VAR_GLOBAL   // PLC tag table "默认变量表"
   "送煤皮带备妥" AT %I0.0 : Bool;
   "送煤皮带运行" AT %I0.1 : Bool;
   "送煤皮带故障" AT %I0.2 : Bool;
   "除铁器备妥" AT %I0.3 : Bool;
   "除铁器运行" AT %I0.4 : Bool;
   "除铁器故障" AT %I0.5 : Bool;
   "定量给煤机备妥" AT %I0.6 : Bool;
   "定量给煤机运行" AT %I0.7 : Bool;
   "定量给煤机故障" AT %I1.0 : Bool;
   "煤粉收尘器备妥" AT %I1.1 : Bool;
   "煤粉收尘器运行" AT %I1.2 : Bool;
   "煤粉收尘器故障" AT %I1.3 : Bool;
   "立磨尾排风机远程" AT %I1.4 : Bool;
   "立磨尾排风机运行" AT %I1.5 : Bool;
   "立磨尾排风机故障" AT %I1.6 : Bool;
   "立磨尾排风机待机" AT %I1.7 : Bool;
   "立磨尾排高压柜远程" AT %I2.0 : Bool;
   "立磨尾排高压柜合闸" AT %I2.1 : Bool;
   "立磨尾排高压柜分闸" AT %I2.2 : Bool;
   "定量给煤机断料信号" AT %I2.3 : Bool;
   "定量给煤机左跑偏信号" AT %I2.4 : Bool;
   "定量给煤机右跑偏信号" AT %I2.5 : Bool;
   "给煤机断链信号" AT %I2.6 : Bool;
   "立磨给煤机累计脉冲" AT %I2.7 : Bool;
   "定量给料机远程" AT %I3.0 : Bool;
   "1#铰刀运行" AT %I3.1 : Bool;
   "2#铰刀运行" AT %I3.2 : Bool;
   "1#分割轮运行" AT %I3.3 : Bool;
   "2#分割轮运行" AT %I3.4 : Bool;
   "3#分割轮运行" AT %I3.5 : Bool;
   "4#分割轮运行" AT %I3.6 : Bool;
   "5#分割轮运行" AT %I3.7 : Bool;
   "立磨主机高压柜远程" AT %I4.0 : Bool;
   "立磨主机高压柜合闸" AT %I4.1 : Bool;
   "立磨主机高压柜分闸" AT %I4.2 : Bool;
   "立磨主机运行" AT %I4.3 : Bool;
   "立磨主机故障" AT %I4.4 : Bool;
   "允许主机启动" AT %I4.5 : Bool;
   "跳停主机" AT %I4.6 : Bool;
   "6#分割轮运行" AT %I5.0 : Bool;
   "7#分割轮运行" AT %I5.1 : Bool;
   "8#分割轮运行" AT %I5.2 : Bool;
   "9#分割轮运行" AT %I5.3 : Bool;
   "10#分割轮运行" AT %I5.4 : Bool;
   "立磨尾排风机水平震动1" AT %IW256 : Int;
   "立磨尾排风机水平震动2" AT %IW258 : Int;
   "立磨尾排风机垂直震动1" AT %IW260 : Int;
   "立磨尾排风机垂直震动2" AT %IW262 : Int;
   "立磨尾排风机入口压力1" AT %IW264 : Int;
   "立磨尾排风机入口压力2" AT %IW266 : Int;
   "立磨尾排风机出口压力1" AT %IW268 : Int;
   "尾排风机入口执行器反馈" AT %IW270 : Int;
   "立磨1#煤粉仓负压" AT %IW272 : Int;
   "立磨2#煤粉仓负压" AT %IW274 : Int;
   "立磨热风管道负压" AT %IW276 : Int;
   "立磨主电机运行电流" AT %IW278 : Int;
   "立磨给煤机流量" AT %IW280 : Int;
   "立磨出口压力1" AT %IW282 : Int;
   "立磨出口压力2" AT %IW284 : Int;
   "立磨尾排风机运行转速" AT %IW288 : Int;
   "立磨尾排风机运行电流" AT %IW290 : Int;
   "立磨尾排风机出口温度1" AT %IW292 : Int;
   "立磨尾排风机入口温度1" AT %IW296 : Int;
   "立磨尾排风机入口温度2" AT %IW298 : Int;
   "立磨入磨口温度" AT %IW300 : Int;
   "1#煤粉仓1#温度" AT %ID304 : DWord;
   "1#煤粉仓2#温度" AT %ID308 : DWord;
   "1#煤粉仓3#温度" AT %ID312 : DWord;
   "1#煤粉仓4#温度" AT %ID316 : DWord;
   "1#煤粉仓5#温度" AT %ID320 : DWord;
   "1#煤粉仓6#温度" AT %ID324 : DWord;
   "2#煤粉仓1#温度" AT %ID328 : DWord;
   "2#煤粉仓2#温度" AT %ID332 : DWord;
   "2#煤粉仓3#温度" AT %ID336 : DWord;
   "2#煤粉仓4#温度" AT %ID340 : DWord;
   "2#煤粉仓5#温度" AT %ID344 : DWord;
   "2#煤粉仓6#温度" AT %ID348 : DWord;
   "立磨机出口温度1" AT %ID352 : DWord;
   "立磨机出口温度2" AT %ID356 : DWord;
   "PID360" AT %ID360 : DWord;
   "PID364" AT %ID364 : DWord;
   "电机绕组U相温度" AT %ID368 : DWord;
   "电机绕组V相温度" AT %ID372 : DWord;
   "电机绕组W相温度" AT %ID376 : DWord;
   "尾排电机前轴温度" AT %ID380 : DWord;
   "尾排电机后轴温度" AT %ID384 : DWord;
   "尾排风机前轴温度" AT %ID388 : DWord;
   "尾排风机后轴温度" AT %ID392 : DWord;
   "PID396" AT %ID396 : DWord;
   "立磨主机远程" AT %I4.7 : Bool;
   "11#分割轮运行" AT %I5.5 : Bool;
   "12#分割轮运行" AT %I5.6 : Bool;
   "立磨主电机轻故障" AT %I5.7 : Bool;
   "1#板式给煤机-褐煤备妥" AT %I6.0 : Bool;
   "1#板式给煤机-褐煤运行" AT %I6.1 : Bool;
   "1#板式给煤机-褐煤故障" AT %I6.2 : Bool;
   "2#板式给煤机-烟煤备妥" AT %I6.3 : Bool;
   "2#板式给煤机-烟煤运行" AT %I6.4 : Bool;
   "2#板式给煤机-烟煤故障" AT %I6.5 : Bool;
   "1#板式给煤机-褐煤脉冲累计" AT %I6.6 : Bool;
   "2#板式给煤机-烟煤脉冲累计" AT %I6.7 : Bool;
   "储气罐阀门远程" AT %I7.0 : Bool;
   "储气罐阀门开到位" AT %I7.1 : Bool;
   "储气罐阀门关到位" AT %I7.2 : Bool;
   "I7_3" AT %I7.3 : Bool;
   "I7_4" AT %I7.4 : Bool;
   "I7_5" AT %I7.5 : Bool;
   "I7_6" AT %I7.6 : Bool;
   "I7_7" AT %I7.7 : Bool;
   "I8_0" AT %I8.0 : Bool;
   "I8_1" AT %I8.1 : Bool;
   "I8_2" AT %I8.2 : Bool;
   "I8_3" AT %I8.3 : Bool;
   "I8_4" AT %I8.4 : Bool;
   "I8_5" AT %I8.5 : Bool;
   "I8_6" AT %I8.6 : Bool;
   "I8_7" AT %I8.7 : Bool;
   "I9_0" AT %I9.0 : Bool;
   "I9_1" AT %I9.1 : Bool;
   "I9_2" AT %I9.2 : Bool;
   "I9_3" AT %I9.3 : Bool;
   "I9_4" AT %I9.4 : Bool;
   "I9_5" AT %I9.5 : Bool;
   "I9_6" AT %I9.6 : Bool;
   "I9_7" AT %I9.7 : Bool;
   "I10_0" AT %I10.0 : Bool;
   "I10_1" AT %I10.1 : Bool;
   "I10_2" AT %I10.2 : Bool;
   "I10_3" AT %I10.3 : Bool;
   "I10_4" AT %I10.4 : Bool;
   "I10_5" AT %I10.5 : Bool;
   "I10_6" AT %I10.6 : Bool;
   "I10_7" AT %I10.7 : Bool;
   "I11_0" AT %I11.0 : Bool;
   "I11_1" AT %I11.1 : Bool;
   "I11_2" AT %I11.2 : Bool;
   "I11_3" AT %I11.3 : Bool;
   "I11_4" AT %I11.4 : Bool;
   "I11_5" AT %I11.5 : Bool;
   "I11_6" AT %I11.6 : Bool;
   "I11_7" AT %I11.7 : Bool;
   "1#板式给煤机-褐煤流量反馈" AT %IW286 : Int;
   "2#板式给煤机-烟煤流量反馈" AT %IW294 : Int;
   "PIW302" AT %IW302 : Int;
   "立磨煤粉仓称重" AT %ID450 : Real;
   "立磨1#煤粉仓称重" AT %ID458 : Real;
   "立磨2#煤粉仓称重" AT %ID466 : Real;
   "PID400" AT %ID400 : DWord;
   "PID404" AT %ID404 : DWord;
   "PID408" AT %ID408 : DWord;
   "PID412" AT %ID412 : DWord;
   "PID416" AT %ID416 : DWord;
   "PID420" AT %ID420 : DWord;
   "PID424" AT %ID424 : DWord;
   "PID428" AT %ID428 : DWord;
   "Tag_22" AT %ID374 : Real;
   "送煤皮带驱动" AT %Q0.0 : Bool;
   "除铁器驱动" AT %Q0.1 : Bool;
   "定量给煤机驱动" AT %Q0.2 : Bool;
   "煤粉收尘器驱动" AT %Q0.3 : Bool;
   "立磨尾排风机停止" AT %Q0.4 : Bool;
   "立磨尾排高压柜合闸驱动" AT %Q0.5 : Bool;
   "立磨尾排风机高压柜分闸" AT %Q0.6 : Bool;
   "立磨尾排风机启动" AT %Q0.7 : Bool;
   "立磨主机高压柜合闸驱动" AT %Q1.0 : Bool;
   "立磨主机高压柜分闸驱动" AT %Q1.1 : Bool;
   "QB4" AT %QB4 : Byte;
   "立磨给煤机流量给定" AT %QW256 : Int;
   "立磨尾排风机转速给定" AT %QW258 : Int;
   "尾排风机入口执行器给定" AT %QW260 : Int;
   "1#板式给煤机-褐煤启停" AT %Q1.2 : Bool;
   "2#板式给煤机-烟煤启停" AT %Q1.3 : Bool;
   "立磨现场皮带报警器" AT %Q1.4 : Bool;
   "立磨中控报警器" AT %Q1.5 : Bool;
   "立磨主机启动" AT %Q1.6 : Bool;
   "立磨主机停止" AT %Q1.7 : Bool;
   "储气罐阀门打开" AT %Q2.0 : Bool;
   "储气罐阀门关闭" AT %Q2.1 : Bool;
   "Q2_2" AT %Q2.2 : Bool;
   "Q2_3" AT %Q2.3 : Bool;
   "Q2_4" AT %Q2.4 : Bool;
   "Q2_5" AT %Q2.5 : Bool;
   "Q2_6" AT %Q2.6 : Bool;
   "Q2_7" AT %Q2.7 : Bool;
   "Q3_0" AT %Q3.0 : Bool;
   "Q3_1" AT %Q3.1 : Bool;
   "Q3_2" AT %Q3.2 : Bool;
   "Q3_3" AT %Q3.3 : Bool;
   "Q3_4" AT %Q3.4 : Bool;
   "Q3_5" AT %Q3.5 : Bool;
   "Q3_6" AT %Q3.6 : Bool;
   "Q3_7" AT %Q3.7 : Bool;
   "1#板式给煤机-褐煤流量给定" AT %QW262 : Int;
   "2#板式给煤机-烟煤流量给定" AT %QW264 : Int;
   "PQW266" AT %QW266 : Int;
   "PQW268" AT %QW268 : Int;
   "PQW270" AT %QW270 : Int;
   "Q4.0" AT %Q4.0 : Bool;
   "Tag_5" AT %M2.0 : Bool;
   "Tag_11" AT %M2.3 : Bool;
   "Tag_19" AT %M2.5 : Bool;
   "Tag_1" AT %MW4 : Word;
   "Tag_8" AT %MW10 : Word;
   "Tag_6" AT %MW12 : Word;
   "Tag_21" AT %MW14 : Word;
   "Tag_16" AT %MW16 : Word;
   "锁风定量给煤机流量累计清零" AT %M30.1 : Bool;
   "Tag_13" AT %MW100 : Word;
   "Tag_12" AT %M300.0 : Bool;
   "Tag_20" AT %M300.1 : Bool;
   "Tag_9" AT %M400.0 : Bool;
   "Tag_17" AT %M400.1 : Bool;
   "1#立磨板式给料流量累计清零" AT %M30.2 : Bool;
   "2#立磨板式给料流量累计清零" AT %M30.3 : Bool;
   "Tag_2" AT %M30.7 : Bool;
   "Tag_80" AT %M80.0 : Bool;
   "Tag_81" AT %M81.0 : Bool;
   "Tag_82" AT %M80.1 : Bool;
   "Tag_83" AT %M80.2 : Bool;
   "Tag_84" AT %M80.3 : Bool;
   "Tag_85" AT %M81.1 : Bool;
   "Clock_Byte" AT %MB0 : Byte;
   "Clock_10Hz" AT %M0.0 : Bool;
   "Clock_5Hz" AT %M0.1 : Bool;
   "Clock_2.5Hz" AT %M0.2 : Bool;
   "Clock_2Hz" AT %M0.3 : Bool;
   "Clock_1.25Hz" AT %M0.4 : Bool;
   "Clock_1Hz" AT %M0.5 : Bool;
   "Clock_0.625Hz" AT %M0.6 : Bool;
   "Clock_0.5Hz" AT %M0.7 : Bool;
   "System_Byte" AT %MB1 : Byte;
   "FirstScan" AT %M1.0 : Bool;
   "DiagStatusUpdate" AT %M1.1 : Bool;
   "AlwaysTRUE" AT %M1.2 : Bool;
   "AlwaysFALSE" AT %M1.3 : Bool;
   "Tag_7" AT %MW200 : Word;
   "Tag_14" AT %MW202 : Word;
   "Tag_15" AT %M200.0 : Bool;
   "Tag_26" AT %M200.1 : Bool;
   "Tag_28" AT %M2.1 : Bool;
   "Tag_29" AT %MW82 : Word;
   "Tag_32" AT %M10.0 : Bool;
   "Tag_33" AT %MD40 : Real;
   "Tag_34" AT %MD44 : Real;
   "Tag_35" AT %MD48 : Real;
   "Tag_36" AT %M60.0 : Bool;
   "HMI_ALARM_RST" AT %M10.1 : Bool;
   "Tag_38" AT %M10.2 : Bool;
   "Tag_3" AT %T100 : Timer;
   "Tag_4" AT %T101 : Timer;
   "Tag_86" AT %T102 : Timer;
   "Tag_10" AT %C1 : Counter;
   "Tag_18" AT %C2 : Counter;
   "Tag_30" AT %C3 : Counter;
   "Tag_31" AT %C4 : Counter;
END_VAR

DATA_BLOCK "qud"   // DB1
{ S7_Optimized_Access := 'FALSE' }
VERSION : 0.1
   VAR
      送煤皮带启动 : Bool;
      送煤皮带停止 : Bool;
      除铁器启动 : Bool;
      除铁器停止 : Bool;
      定量给煤机启动 : Bool;
      定量给煤机停止 : Bool;
      煤粉收尘器启动 : Bool;
      煤粉收尘器停止 : Bool;
      STAT8 : Bool;
      STAT9 : Bool;
      立磨主机高压柜合闸 : Bool;
      立磨主机高压柜分闸 : Bool;
      立磨尾排风机启动 : Bool;
      立磨尾排风机停止 : Bool;
      立磨尾排高压柜合闸 : Bool;
      立磨尾排高压柜分闸 : Bool;
      "1#立磨板式给料机启动" : Bool;
      "1#立磨板式给料机停止" : Bool;
      "2#立磨板式给料机启动" : Bool;
      "2#立磨板式给料机停止" : Bool;
      储气罐气源阀门打开 : Bool;
      储气罐气源阀门关闭 : Bool;
      立磨主机启动 : Bool;
      立磨主机停止 : Bool;
   END_VAR
BEGIN
END_DATA_BLOCK

DATA_BLOCK "MNL"   // DB2
{ S7_Optimized_Access := 'FALSE' }
VERSION : 0.1
   VAR
      锁风定量给煤机 : Real := 44.0;
      锁风定量给煤机流量反馈 : Real;
      立磨尾排水平振动1 : Real;
      立磨尾排水平振动2 : Real;
      立磨尾排风机垂直振动1 : Real;
      立磨尾排风机垂直振动2 : Real;
      立磨尾排风机出口压力1 : Real;
      立磨尾排风机出口压力2 : Real;
      STAT8 : Real := 56.07639;
      立磨尾排风机出口温度2 : Real;
      STAT10 : Real := 47.39583;
      STAT11 : Real := 46.52778;
      立磨尾排风机入口压力1 : Real := -2147.512;
      立磨尾排风机入口压力2 : Real := -2461.689;
      "立磨1#煤粉仓负压" : Real := -300.0;
      "立磨2#煤粉仓负压" : Real := -272.9167;
      立磨热风管道负压 : Real := -562.5;
      立磨煤粉仓称重 : Real := 101.51;
      "立磨1#煤粉仓称重" : Real := 8.44;
      "立磨2#煤粉仓称重" : Real := 13.24;
      尾排风机运行频率 : Real := 744.2824;
      尾排风机运行电流 : Real := 41.25;
      主电机运行电流 : Real;
      立磨尾排风机转速给定 : Real := 500.0;
      锁风定量给煤机流量累计 : Real := 30006.97;
      "1#煤粉仓1#温度" : Real := 37.0;
      "1#煤粉仓2#温度" : Real := 36.0;
      "1#煤粉仓3#温度" : Real := 37.0;
      "1#煤粉仓4#温度" : Real := 36.0;
      "1#煤粉仓5#温度" : Real := 36.0;
      "1#煤粉仓6#温度" : Real := 37.0;
      "2#煤粉仓1#温度" : Real := 37.0;
      "2#煤粉仓2#温度" : Real := 36.0;
      "2#煤粉仓3#温度" : Real := 37.0;
      "2#煤粉仓4#温度" : Real := 37.0;
      "2#煤粉仓5#温度" : Real := 37.0;
      "2#煤粉仓6#温度" : Real := 37.0;
      电机绕组U相温度 : Real := 59.0;
      电机绕组V相温度 : Real := 57.0;
      电机绕组W相温度 : Real := 59.0;
      尾排电机前轴温度 : Real := 34.0;
      尾排电机后轴温度 : Real := 40.0;
      尾排风机前轴温度 : Real := 144.8206;
      尾排风机后轴温度 : Real;
      立磨机出口温度1 : Real;
      立磨机出口温度2 : Real := 43.0;
      STAT46 : Real := 46.0;
      STAT47 : Real := 62.0;
      STAT48 : Real := 58.0;
      立磨尾排风机出口温度1 : Real := -1753.472;
      立磨尾排风机入口温度1 : Real := -1707.176;
      立磨尾排风机入口温度2 : Real;
      尾排风机执行器开度给定 : Real;
      尾排风机执行器开度反馈 : Real;
      立磨机出口压力1 : Real;
      立磨机出口压力2 : Real;
      立磨主电机入磨口温度 : Real;
      "1#立磨板式给料反馈" : Real;
      "2#立磨板式给料反馈" : Real;
      "1#立磨板式给料给定" : Real;
      "2#立磨板式给料给定" : Real;
      "1#立磨板式给料累计" : Real;
      "2#立磨板式给料累计" : Real;
      STAT63 : Real;
      STAT64 : Real;
      STAT65 : Real;
   END_VAR
BEGIN
END_DATA_BLOCK

DATA_BLOCK "TIMEDB"   // DB3
{ S7_Optimized_Access := 'TRUE' }
VERSION : 0.1
   VAR
      T1 : IEC_TIMER;
      T2 : IEC_TIMER;
      T3 : IEC_TIMER;
      T4 : IEC_TIMER;
      T5 : IEC_TIMER;
      T6 : IEC_TIMER;
      T7 : IEC_TIMER;
      T8 : IEC_TIMER;
      T9 : IEC_TIMER;
      T10 : IEC_TIMER;
      T11 : IEC_TIMER;
      T12 : IEC_TIMER;
      T13 : IEC_TIMER;
      T14 : IEC_TIMER;
      T15 : IEC_TIMER;
      T16 : IEC_TIMER;
      T17 : IEC_TIMER;
      T18 : IEC_TIMER;
      T19 : IEC_TIMER;
      T20 : IEC_TIMER;
      T21 : IEC_TIMER;
      T22 : IEC_TIMER;
      T23 : IEC_TIMER;
      T24 : IEC_TIMER;
      T25 : IEC_TIMER;
      T26 : IEC_TIMER;
      T27 : IEC_TIMER;
      T28 : IEC_TIMER;
      T29 : IEC_TIMER;
      T30 : IEC_TIMER;
      T31 : IEC_TIMER;
      T32 : IEC_TIMER;
      T33 : IEC_TIMER;
      T34 : IEC_TIMER;
      T35 : IEC_TIMER;
      T36 : IEC_TIMER;
      T37 : IEC_TIMER;
      T38 : IEC_TIMER;
      T39 : IEC_TIMER;
      T40 : IEC_TIMER;
      T41 : IEC_TIMER;
      T42 : IEC_TIMER;
      T43 : IEC_TIMER;
      T44 : IEC_TIMER;
      T45 : IEC_TIMER;
      T46 : IEC_TIMER;
      T47 : IEC_TIMER;
      T48 : IEC_TIMER;
      T49 : IEC_TIMER;
      T50 : IEC_TIMER;
      T51 : IEC_TIMER;
      T52 : IEC_TIMER;
      T53 : IEC_TIMER;
      T54 : IEC_TIMER;
      T55 : IEC_TIMER;
      T56 : IEC_TIMER;
      T57 : IEC_TIMER;
      T58 : IEC_TIMER;
      T59 : IEC_TIMER;
      T60 : IEC_TIMER;
      T61 : IEC_TIMER;
      T62 : IEC_TIMER;
      T63 : IEC_TIMER;
      T64 : IEC_TIMER;
      T65 : IEC_TIMER;
      T66 : IEC_TIMER;
      T67 : IEC_TIMER;
      T68 : IEC_TIMER;
      T69 : IEC_TIMER;
      T70 : IEC_TIMER;
      T71 : IEC_TIMER;
      T72 : IEC_TIMER;
      T73 : IEC_TIMER;
      T74 : IEC_TIMER;
      T75 : IEC_TIMER;
      T76 : IEC_TIMER;
      T77 : IEC_TIMER;
      T78 : IEC_TIMER;
      T79 : IEC_TIMER;
      T80 : IEC_TIMER;
      T81 : IEC_TIMER;
      T82 : IEC_TIMER;
      T83 : IEC_TIMER;
      T84 : IEC_TIMER;
      T85 : IEC_TIMER;
      T86 : IEC_TIMER;
      T87 : IEC_TIMER;
      T88 : IEC_TIMER;
      T89 : IEC_TIMER;
      T90 : IEC_TIMER;
      T91 : IEC_TIMER;
      T92 : IEC_TIMER;
      T93 : IEC_TIMER;
      T94 : IEC_TIMER;
      T95 : IEC_TIMER;
      T96 : IEC_TIMER;
      T97 : IEC_TIMER;
      T98 : IEC_TIMER;
      T99 : IEC_TIMER;
      T100 : IEC_TIMER;
   END_VAR
BEGIN
END_DATA_BLOCK

DATA_BLOCK "累计功能块_DB_1"   // DB4
{ S7_Optimized_Access := 'FALSE' }
VERSION : 0.1
// stored: InstanceOfName 累计功能块
"累计功能块"
BEGIN
END_DATA_BLOCK

DATA_BLOCK "累计功能块_DB"   // DB5
{ S7_Optimized_Access := 'FALSE' }
VERSION : 0.1
// stored: InstanceOfName 累计功能块
"累计功能块"
BEGIN
END_DATA_BLOCK

DATA_BLOCK "累计功能块_DB_2"   // DB6
{ S7_Optimized_Access := 'FALSE' }
VERSION : 0.1
// stored: InstanceOfName 累计功能块
"累计功能块"
BEGIN
END_DATA_BLOCK

DATA_BLOCK "DB9_P"   // DB9
{ S7_Optimized_Access := 'FALSE' }
VERSION : 0.1
   VAR
      P1 : Bool;
      P2 : Bool;
      P3 : Bool;
      P4 : Bool;
      P5 : Bool;
      P6 : Bool;
      P7 : Bool;
      P8 : Bool;
      P9 : Bool;
      P10 : Bool;
      P11 : Bool;
      P12 : Bool;
      P13 : Bool;
      P14 : Bool;
      P15 : Bool;
      P16 : Bool;
      P17 : Bool;
      P18 : Bool;
      P19 : Bool;
      P20 : Bool;
      P21 : Bool;
      P22 : Bool;
      P23 : Bool;
      P24 : Bool;
      P25 : Bool;
      P26 : Bool;
      P27 : Bool;
      P28 : Bool;
      P29 : Bool;
      P30 : Bool;
      P31 : Bool;
      P32 : Bool;
      P33 : Bool;
      P34 : Bool;
      P35 : Bool;
      P36 : Bool;
      P37 : Bool;
      P38 : Bool;
      P39 : Bool;
      P40 : Bool;
      P41 : Bool;
      P42 : Bool;
      P43 : Bool;
      P44 : Bool;
      P45 : Bool;
      P46 : Bool;
      P47 : Bool;
      P48 : Bool;
      P49 : Bool;
      P50 : Bool;
      P51 : Bool;
      P52 : Bool;
      P53 : Bool;
      P54 : Bool;
      P55 : Bool;
      P56 : Bool;
      P57 : Bool;
      P58 : Bool;
      P59 : Bool;
      P60 : Bool;
      P61 : Bool;
      P62 : Bool;
      P63 : Bool;
      P64 : Bool;
      P65 : Bool;
      P66 : Bool;
      P67 : Bool;
      P68 : Bool;
      P69 : Bool;
      P70 : Bool;
      P71 : Bool;
      P72 : Bool;
      P73 : Bool;
      P74 : Bool;
      P75 : Bool;
      P76 : Bool;
      P77 : Bool;
      P78 : Bool;
      P79 : Bool;
      P80 : Bool;
      P81 : Bool;
      P82 : Bool;
      P83 : Bool;
      P84 : Bool;
      P85 : Bool;
      P86 : Bool;
      P87 : Bool;
      P88 : Bool;
      P89 : Bool;
      P90 : Bool;
      P91 : Bool;
      P92 : Bool;
      P93 : Bool;
   END_VAR
BEGIN
END_DATA_BLOCK

DATA_BLOCK "FB11_DATA_ALARM_FB_DB"   // DB11
{ S7_Optimized_Access := 'FALSE' }
VERSION : 0.1
// stored: InstanceOfName FB11_DATA_ALARM_FB
"FB11_DATA_ALARM_FB"
BEGIN
END_DATA_BLOCK

FUNCTION_BLOCK "累计功能块"   // FB1, LAD
{ S7_Optimized_Access := 'FALSE' }
VERSION : 0.1
   VAR_INPUT
      CLEAR : Bool;   // 清零
      IN : Bool;   // 累计脉冲信号
   END_VAR
   VAR_OUTPUT
      OUT1 : Real;
   END_VAR
   VAR
      STAT2 : Real;
      STAT3 : Real;
      STAT4 : Real;
      P1 : Bool;
   END_VAR
   VAR_TEMP   // added for the SCL form of the ladder/FBD networks
      _w1 : Bool;
   END_VAR
BEGIN

REGION Network 1
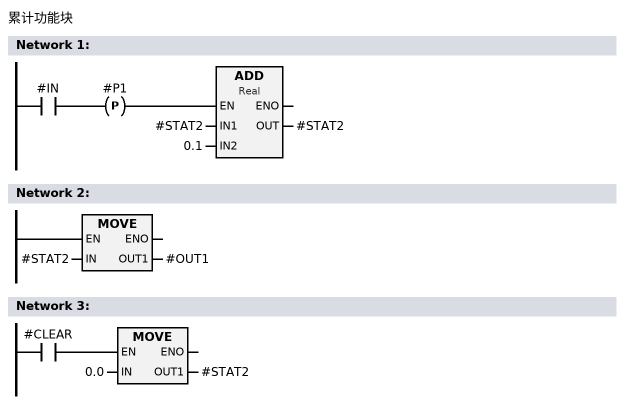
   RUNG wire#powerrail
      Contact( #IN )
      P_Trig( #P1 )
      { S7_Templates := "SrcType := Real"; S7_GenerateENO := "TRUE" } Add(in1 := #STAT2, in2 := 0.1, out => #STAT2)
   END_RUNG
   // the same network as SCL:
   #_w1 := #IN AND NOT #P1;   // rising edge
   #P1 := #IN;
   IF #_w1 THEN #STAT2 := #STAT2 + 0.1; END_IF;
END_REGION

REGION Network 2
   RUNG wire#powerrail
      { S7_GenerateENO := "TRUE" } Move(in := #STAT2, out1 => #OUT1)
   END_RUNG
   // the same network as SCL:
   #OUT1 := #STAT2;
END_REGION

REGION Network 3
   RUNG wire#powerrail
      Contact( #CLEAR )
      { S7_GenerateENO := "TRUE" } Move(in := 0.0, out1 => #STAT2)
   END_RUNG
   // the same network as SCL:
   IF #CLEAR THEN #STAT2 := 0.0; END_IF;
END_REGION
END_FUNCTION_BLOCK

FUNCTION_BLOCK "FB11_DATA_ALARM_FB"   // FB11, LAD
{ S7_Optimized_Access := 'FALSE' }
VERSION : 0.1
   VAR
      PIW256 : "FB330_DATA_ALARM";
      PIW258 : "FB330_DATA_ALARM";
      PIW260 : "FB330_DATA_ALARM";
      PIW262 : "FB330_DATA_ALARM";
      PIW264 : "FB330_DATA_ALARM";
      PIW266 : "FB330_DATA_ALARM";
      PIW268 : "FB330_DATA_ALARM";
      PIW270 : "FB330_DATA_ALARM";
      PIW272 : "FB330_DATA_ALARM";
      PIW274 : "FB330_DATA_ALARM";
      PIW276 : "FB330_DATA_ALARM";
      PIW278 : "FB330_DATA_ALARM";
      PIW280 : "FB330_DATA_ALARM";
      PIW282 : "FB330_DATA_ALARM";
      PIW284 : "FB330_DATA_ALARM";
      PIW286 : "FB330_DATA_ALARM";
      PIW288 : "FB330_DATA_ALARM";
      PIW290 : "FB330_DATA_ALARM";
      PIW292 : "FB330_DATA_ALARM";
      PIW294 : "FB330_DATA_ALARM";
      PIW296 : "FB330_DATA_ALARM";
      PIW298 : "FB330_DATA_ALARM";
      PIW300 : "FB330_DATA_ALARM";
      PIW302 : "FB330_DATA_ALARM";
      PID304 : "FB330_DATA_ALARM";
      PID308 : "FB330_DATA_ALARM";
      PID312 : "FB330_DATA_ALARM";
      PID316 : "FB330_DATA_ALARM";
      PID320 : "FB330_DATA_ALARM";
      PID324 : "FB330_DATA_ALARM";
      PID328 : "FB330_DATA_ALARM";
      PID332 : "FB330_DATA_ALARM";
      PID336 : "FB330_DATA_ALARM";
      PID340 : "FB330_DATA_ALARM";
      PID344 : "FB330_DATA_ALARM";
      PID348 : "FB330_DATA_ALARM";
      PID352 : "FB330_DATA_ALARM";
      PID356 : "FB330_DATA_ALARM";
      PID360 : "FB330_DATA_ALARM";
      PID364 : "FB330_DATA_ALARM";
      PID368 : "FB330_DATA_ALARM";
      PID372 : "FB330_DATA_ALARM";
      PID376 : "FB330_DATA_ALARM";
      PID380 : "FB330_DATA_ALARM";
      PID384 : "FB330_DATA_ALARM";
      PID388 : "FB330_DATA_ALARM";
      PID392 : "FB330_DATA_ALARM";
      PID396 : "FB330_DATA_ALARM";
      IW110 : "FB330_DATA_ALARM";
      IW112 : "FB330_DATA_ALARM";
      IW114 : "FB330_DATA_ALARM";
      IW116 : "FB330_DATA_ALARM";
      PID400 : "FB330_DATA_ALARM";
      PID408 : "FB330_DATA_ALARM";
      PID416 : "FB330_DATA_ALARM";
      Static4 : "FB330_DATA_ALARM";
      Static5 : "FB330_DATA_ALARM";
      Static6 : "FB330_DATA_ALARM";
      Static7 : "FB330_DATA_ALARM";
      Static8 : "FB330_DATA_ALARM";
      Static9 : "FB330_DATA_ALARM";
      Static10 : "FB330_DATA_ALARM";
   END_VAR
BEGIN

REGION Network 1
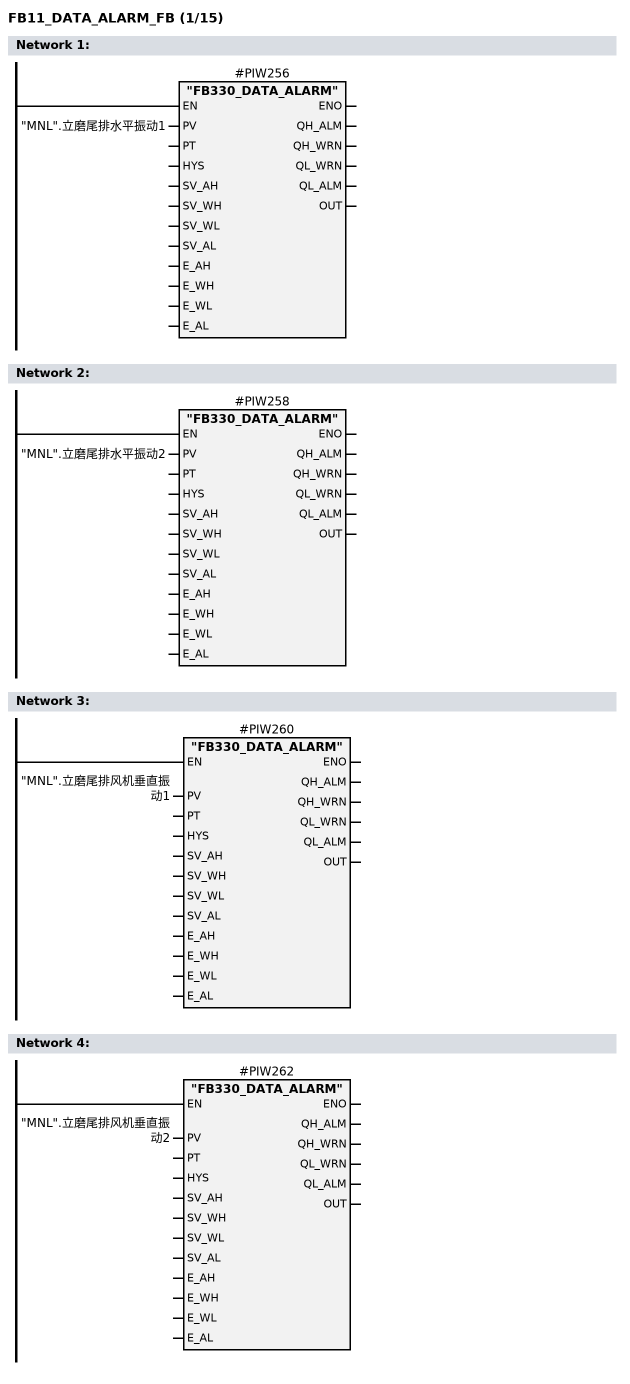
   RUNG wire#powerrail
      #PIW256(PV := "MNL".立磨尾排水平振动1, PT :=, HYS :=, SV_AH :=, SV_WH :=, SV_WL :=, SV_AL :=, E_AH :=, E_WH :=, E_WL :=, E_AL :=, QH_ALM =>, QH_WRN =>, QL_WRN =>, QL_ALM =>, OUT =>)
   END_RUNG
   // the same network as SCL:
   #PIW256(PV := "MNL".立磨尾排水平振动1);   // "FB330_DATA_ALARM"
END_REGION

REGION Network 2
   RUNG wire#powerrail
      #PIW258(PV := "MNL".立磨尾排水平振动2, PT :=, HYS :=, SV_AH :=, SV_WH :=, SV_WL :=, SV_AL :=, E_AH :=, E_WH :=, E_WL :=, E_AL :=, QH_ALM =>, QH_WRN =>, QL_WRN =>, QL_ALM =>, OUT =>)
   END_RUNG
   // the same network as SCL:
   #PIW258(PV := "MNL".立磨尾排水平振动2);   // "FB330_DATA_ALARM"
END_REGION

REGION Network 3
   RUNG wire#powerrail
      #PIW260(PV := "MNL".立磨尾排风机垂直振动1, PT :=, HYS :=, SV_AH :=, SV_WH :=, SV_WL :=, SV_AL :=, E_AH :=, E_WH :=, E_WL :=, E_AL :=, QH_ALM =>, QH_WRN =>, QL_WRN =>, QL_ALM =>, OUT =>)
   END_RUNG
   // the same network as SCL:
   #PIW260(PV := "MNL".立磨尾排风机垂直振动1);   // "FB330_DATA_ALARM"
END_REGION

REGION Network 4
   RUNG wire#powerrail
      #PIW262(PV := "MNL".立磨尾排风机垂直振动2, PT :=, HYS :=, SV_AH :=, SV_WH :=, SV_WL :=, SV_AL :=, E_AH :=, E_WH :=, E_WL :=, E_AL :=, QH_ALM =>, QH_WRN =>, QL_WRN =>, QL_ALM =>, OUT =>)
   END_RUNG
   // the same network as SCL:
   #PIW262(PV := "MNL".立磨尾排风机垂直振动2);   // "FB330_DATA_ALARM"
END_REGION

REGION Network 5
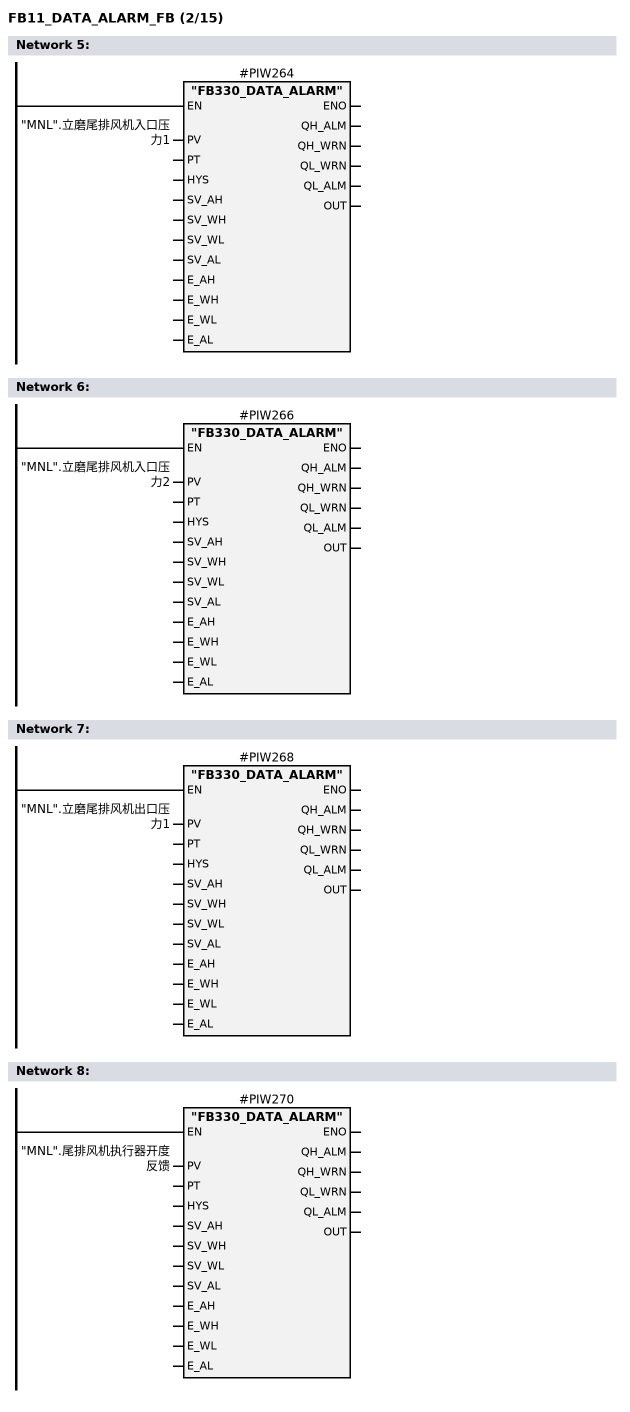
   RUNG wire#powerrail
      #PIW264(PV := "MNL".立磨尾排风机入口压力1, PT :=, HYS :=, SV_AH :=, SV_WH :=, SV_WL :=, SV_AL :=, E_AH :=, E_WH :=, E_WL :=, E_AL :=, QH_ALM =>, QH_WRN =>, QL_WRN =>, QL_ALM =>, OUT =>)
   END_RUNG
   // the same network as SCL:
   #PIW264(PV := "MNL".立磨尾排风机入口压力1);   // "FB330_DATA_ALARM"
END_REGION

REGION Network 6
   RUNG wire#powerrail
      #PIW266(PV := "MNL".立磨尾排风机入口压力2, PT :=, HYS :=, SV_AH :=, SV_WH :=, SV_WL :=, SV_AL :=, E_AH :=, E_WH :=, E_WL :=, E_AL :=, QH_ALM =>, QH_WRN =>, QL_WRN =>, QL_ALM =>, OUT =>)
   END_RUNG
   // the same network as SCL:
   #PIW266(PV := "MNL".立磨尾排风机入口压力2);   // "FB330_DATA_ALARM"
END_REGION

REGION Network 7
   RUNG wire#powerrail
      #PIW268(PV := "MNL".立磨尾排风机出口压力1, PT :=, HYS :=, SV_AH :=, SV_WH :=, SV_WL :=, SV_AL :=, E_AH :=, E_WH :=, E_WL :=, E_AL :=, QH_ALM =>, QH_WRN =>, QL_WRN =>, QL_ALM =>, OUT =>)
   END_RUNG
   // the same network as SCL:
   #PIW268(PV := "MNL".立磨尾排风机出口压力1);   // "FB330_DATA_ALARM"
END_REGION

REGION Network 8
   RUNG wire#powerrail
      #PIW270(PV := "MNL".尾排风机执行器开度反馈, PT :=, HYS :=, SV_AH :=, SV_WH :=, SV_WL :=, SV_AL :=, E_AH :=, E_WH :=, E_WL :=, E_AL :=, QH_ALM =>, QH_WRN =>, QL_WRN =>, QL_ALM =>, OUT =>)
   END_RUNG
   // the same network as SCL:
   #PIW270(PV := "MNL".尾排风机执行器开度反馈);   // "FB330_DATA_ALARM"
END_REGION

REGION Network 9
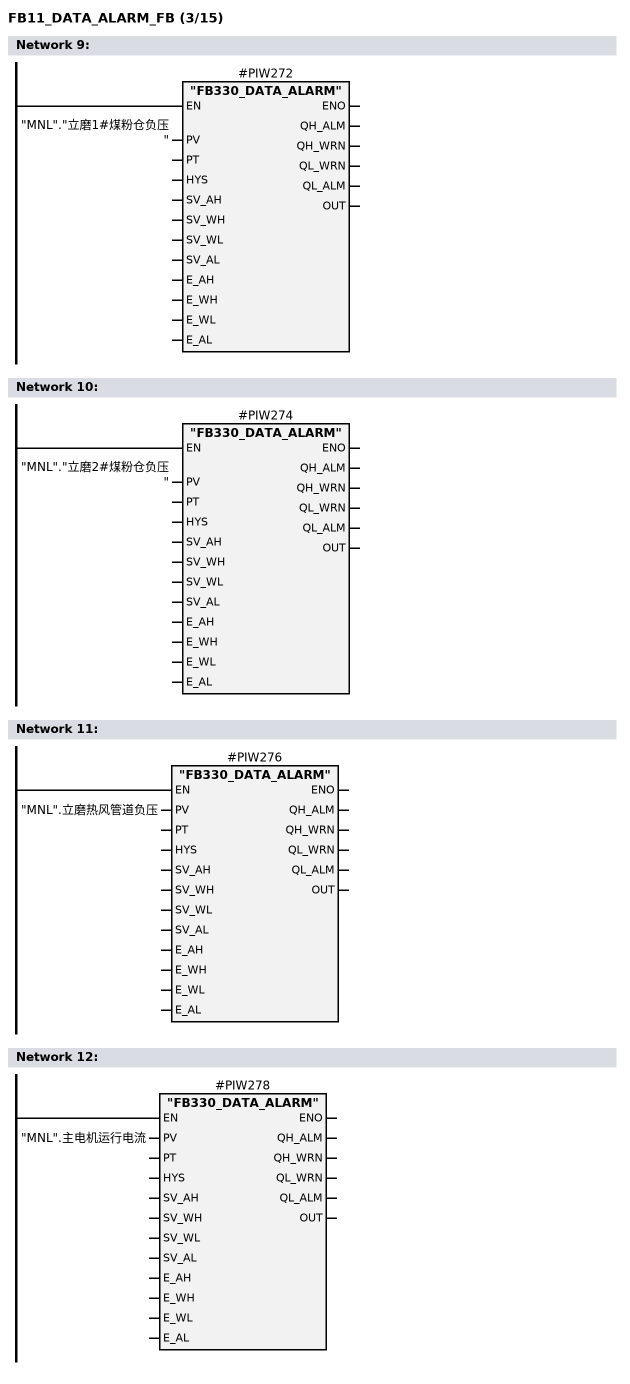
   RUNG wire#powerrail
      #PIW272(PV := "MNL"."立磨1#煤粉仓负压", PT :=, HYS :=, SV_AH :=, SV_WH :=, SV_WL :=, SV_AL :=, E_AH :=, E_WH :=, E_WL :=, E_AL :=, QH_ALM =>, QH_WRN =>, QL_WRN =>, QL_ALM =>, OUT =>)
   END_RUNG
   // the same network as SCL:
   #PIW272(PV := "MNL"."立磨1#煤粉仓负压");   // "FB330_DATA_ALARM"
END_REGION

REGION Network 10
   RUNG wire#powerrail
      #PIW274(PV := "MNL"."立磨2#煤粉仓负压", PT :=, HYS :=, SV_AH :=, SV_WH :=, SV_WL :=, SV_AL :=, E_AH :=, E_WH :=, E_WL :=, E_AL :=, QH_ALM =>, QH_WRN =>, QL_WRN =>, QL_ALM =>, OUT =>)
   END_RUNG
   // the same network as SCL:
   #PIW274(PV := "MNL"."立磨2#煤粉仓负压");   // "FB330_DATA_ALARM"
END_REGION

REGION Network 11
   RUNG wire#powerrail
      #PIW276(PV := "MNL".立磨热风管道负压, PT :=, HYS :=, SV_AH :=, SV_WH :=, SV_WL :=, SV_AL :=, E_AH :=, E_WH :=, E_WL :=, E_AL :=, QH_ALM =>, QH_WRN =>, QL_WRN =>, QL_ALM =>, OUT =>)
   END_RUNG
   // the same network as SCL:
   #PIW276(PV := "MNL".立磨热风管道负压);   // "FB330_DATA_ALARM"
END_REGION

REGION Network 12
   RUNG wire#powerrail
      #PIW278(PV := "MNL".主电机运行电流, PT :=, HYS :=, SV_AH :=, SV_WH :=, SV_WL :=, SV_AL :=, E_AH :=, E_WH :=, E_WL :=, E_AL :=, QH_ALM =>, QH_WRN =>, QL_WRN =>, QL_ALM =>, OUT =>)
   END_RUNG
   // the same network as SCL:
   #PIW278(PV := "MNL".主电机运行电流);   // "FB330_DATA_ALARM"
END_REGION

REGION Network 13
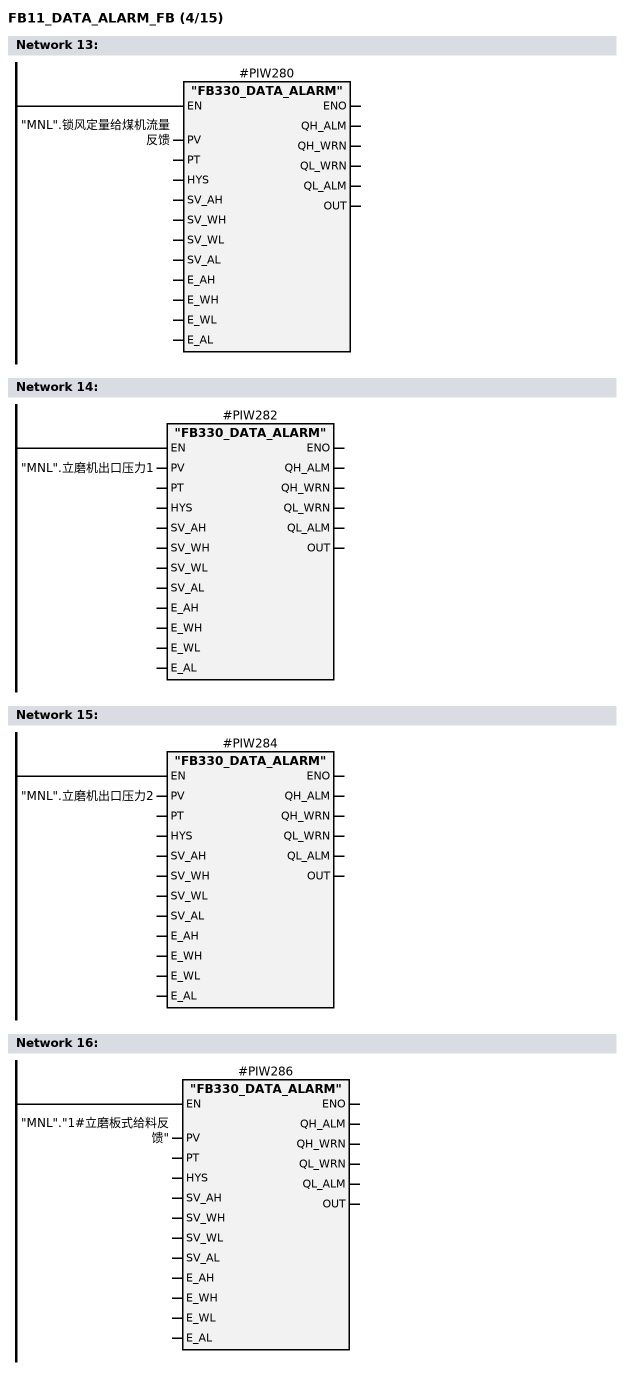
   RUNG wire#powerrail
      #PIW280(PV := "MNL".锁风定量给煤机流量反馈, PT :=, HYS :=, SV_AH :=, SV_WH :=, SV_WL :=, SV_AL :=, E_AH :=, E_WH :=, E_WL :=, E_AL :=, QH_ALM =>, QH_WRN =>, QL_WRN =>, QL_ALM =>, OUT =>)
   END_RUNG
   // the same network as SCL:
   #PIW280(PV := "MNL".锁风定量给煤机流量反馈);   // "FB330_DATA_ALARM"
END_REGION

REGION Network 14
   RUNG wire#powerrail
      #PIW282(PV := "MNL".立磨机出口压力1, PT :=, HYS :=, SV_AH :=, SV_WH :=, SV_WL :=, SV_AL :=, E_AH :=, E_WH :=, E_WL :=, E_AL :=, QH_ALM =>, QH_WRN =>, QL_WRN =>, QL_ALM =>, OUT =>)
   END_RUNG
   // the same network as SCL:
   #PIW282(PV := "MNL".立磨机出口压力1);   // "FB330_DATA_ALARM"
END_REGION

REGION Network 15
   RUNG wire#powerrail
      #PIW284(PV := "MNL".立磨机出口压力2, PT :=, HYS :=, SV_AH :=, SV_WH :=, SV_WL :=, SV_AL :=, E_AH :=, E_WH :=, E_WL :=, E_AL :=, QH_ALM =>, QH_WRN =>, QL_WRN =>, QL_ALM =>, OUT =>)
   END_RUNG
   // the same network as SCL:
   #PIW284(PV := "MNL".立磨机出口压力2);   // "FB330_DATA_ALARM"
END_REGION

REGION Network 16
   RUNG wire#powerrail
      #PIW286(PV := "MNL"."1#立磨板式给料反馈", PT :=, HYS :=, SV_AH :=, SV_WH :=, SV_WL :=, SV_AL :=, E_AH :=, E_WH :=, E_WL :=, E_AL :=, QH_ALM =>, QH_WRN =>, QL_WRN =>, QL_ALM =>, OUT =>)
   END_RUNG
   // the same network as SCL:
   #PIW286(PV := "MNL"."1#立磨板式给料反馈");   // "FB330_DATA_ALARM"
END_REGION

REGION Network 17